(* Logix 5000 project; controller MV vendor 1 type 14 code 217 rev 31.11; software revision 31.00; part 28 of 53 *)
(* tags used below, declared in another part *)
   active : BOOL;
   CWD : CHECKWORD_FLAGS;
   FVHR18_2505 : PlantItem;   // Valve FVHR18_25/05
   FVHR18_2506 : PlantItem;   // Valve FVHR18_25/06
   FVHR26_3101 : PlantItem;   // Valve FVHR26_31/01
   FVHR26_3102 : PlantItem;   // Valve FVHR26_31/02
   FVHR26_3103 : PlantItem;   // Valve FVHR26_31/03
   FVHRCH201 : PlantItem;   // Valve FVHRCH201
   FVHRCH202 : PlantItem;   // Valve FVHRCH202
   FVHRCW01 : PlantItem;   // Valve FVHRCW01
   FVHRM01 : PlantItem;   // Valve FVHRM01
   FVHRM02 : PlantItem;   // Valve FVHRM02
   FVHRM03 : PlantItem;   // Valve FVHRM03
   FVHRM04 : PlantItem;   // Valve FVHRM04
   FVHRMD01 : PlantItem;   // Valve FVHRMD01
   IGI_TestBit : BOOL;
   MC_B243 : INT[255];   // CH2 ROUTE Channel 2 route requ est flags
   MC_CD_T1 : PlantItem;   // CD_T1
   MC_CH2_CIP_BYPASS_Conditions : BOOL;
   MC_CH2_CIP_BYPASS_DrainConditions : BOOL;
   MC_CH2_CIP_Messages : STRING[20];   // CH2 CIP Scada Messages
   MC_CH2_CIP_YST_Scb_Bypass : BOOL;
   MC_CH2_FVBYPASS_H2O_Flush : BOOL;
   MC_CIP_CH2_Strings_HopRinse : STRING[30];
   MC_CIP_String_Result : DINT;
   MC_FL_D1 : PlantItem;   // FL_D1
   MC_N10 : INT[255];   // SETTINGS
   MC_N100 : INT[255];   // C1_PLC Channel 1 PLC data
   MC_N104 : INT[255];   // CH1 REPORT Channel 1 CIP report file
   MC_N120 : INT[255];   // C2 PLC Channel 2 PLC data
   MC_N122 : INT[255];   // CH2 PROG Channel 2 CIP progra m
   MC_N124 : INT[255];   // CH2 REPORT Channel 2 CIP report file
   MC_N200 : INT[255];   // CHK_WORK Plant item fault che cking work area
   MC_N7 : INT[255];   // INTEGER
   MC_N80 : INT[255];   // SRV1_PLC Detergent tank 1 ser vice PLC data
   MC_N80_19_0_Storagebit : BOOL;
   MC_N81 : INT[255];   // SV1_PC Detergent tank 1 ser vice PC to PLC data
   MC_P3 : PlantItem;   // P3
   MC_SFile : INT[255];   // SLC Equivalent System File, So Original Code Can Remain
   MC_SV1 : PlantItem;   // SV1
   MC_T125 : TIMER[255];   // CH2 TIMERS Channel 2 timers
   MC_T4 : TIMER[255];   // TIMER
   MC_T85 : TIMER[255];   // SV1 TIMERS Detergent tank 1 ser vice timers
(* MC_Common, continued *)

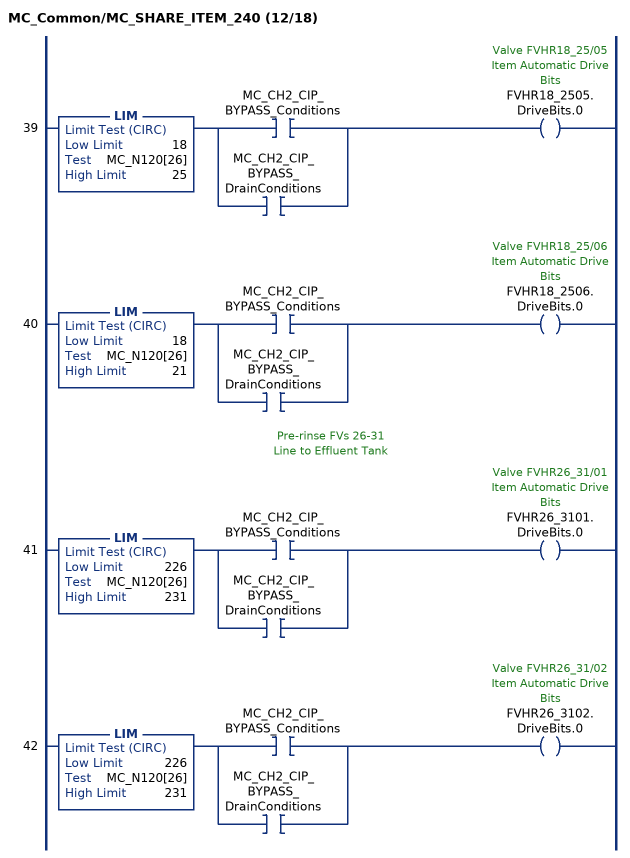
   [picture p556: MC_Common/MC_SHARE_ITEM_240 rungs 39-42]
   39: LIM(18,MC_N120[26],25)[XIC(MC_CH2_CIP_BYPASS_Conditions) ,XIC(MC_CH2_CIP_BYPASS_DrainConditions) ]OTE(FVHR18_2505.DriveBits.0);
   40: LIM(18,MC_N120[26],21)[XIC(MC_CH2_CIP_BYPASS_Conditions) ,XIC(MC_CH2_CIP_BYPASS_DrainConditions) ]OTE(FVHR18_2506.DriveBits.0);
   // Pre-rinse FVs 26-31
   // Line to Effluent Tank
   41: LIM(226,MC_N120[26],231)[XIC(MC_CH2_CIP_BYPASS_Conditions) ,XIC(MC_CH2_CIP_BYPASS_DrainConditions) ]OTE(FVHR26_3101.DriveBits.0);
   42: LIM(226,MC_N120[26],231)[XIC(MC_CH2_CIP_BYPASS_Conditions) ,XIC(MC_CH2_CIP_BYPASS_DrainConditions) ]OTE(FVHR26_3102.DriveBits.0);
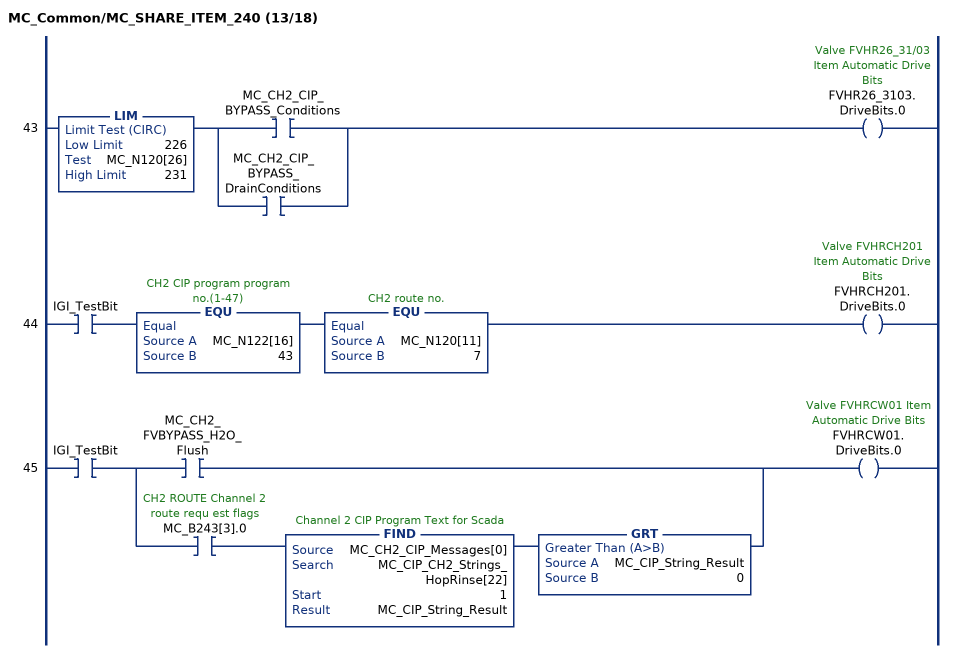
   43: LIM(226,MC_N120[26],231)[XIC(MC_CH2_CIP_BYPASS_Conditions) ,XIC(MC_CH2_CIP_BYPASS_DrainConditions) ]OTE(FVHR26_3103.DriveBits.0);
   44: XIC(IGI_TestBit)EQU(MC_N122[16],43)EQU(MC_N120[11],7)OTE(FVHRCH201.DriveBits.0);
   45: XIC(IGI_TestBit)[XIC(MC_CH2_FVBYPASS_H2O_Flush) ,XIC(MC_B243[3].0) FIND(MC_CH2_CIP_Messages[0],MC_CIP_CH2_Strings_HopRinse[22],1,MC_CIP_String_Result) GRT(MC_CIP_String_Result,0) ]OTE(FVHRCW01.DriveBits.0);
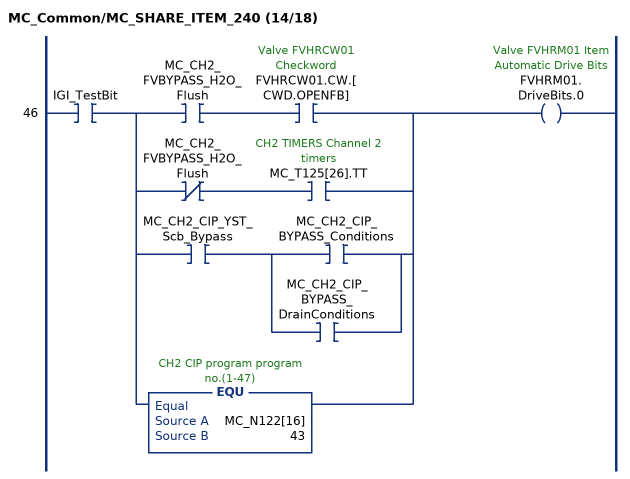
   46: XIC(IGI_TestBit)[XIC(MC_CH2_FVBYPASS_H2O_Flush) XIC(FVHRCW01.CW.[CWD.OPENFB]) ,XIO(MC_CH2_FVBYPASS_H2O_Flush) XIC(MC_T125[26].TT) ,XIC(MC_CH2_CIP_YST_Scb_Bypass) [XIC(MC_CH2_CIP_BYPASS_Conditions) ,XIC(MC_CH2_CIP_BYPASS_DrainConditions) ] ,EQU(MC_N122[16],43) ]OTE(FVHRM01.DriveBits.0);
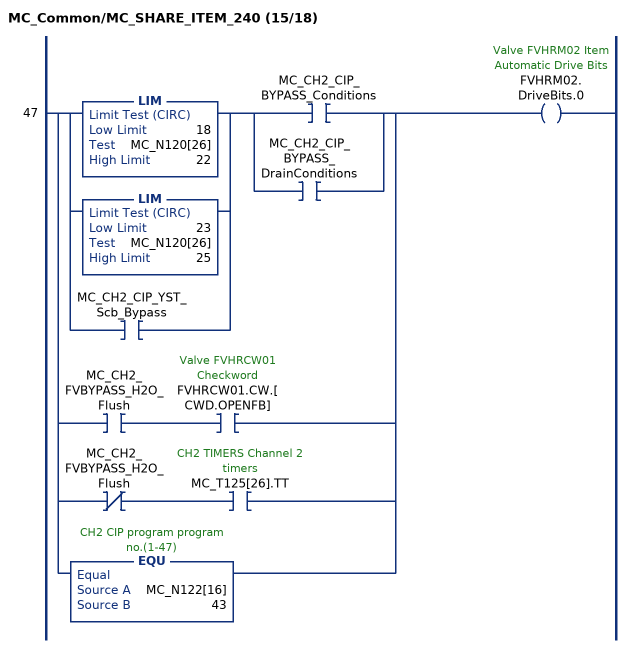
   47: [[LIM(18,MC_N120[26],22) ,LIM(23,MC_N120[26],25) ,XIC(MC_CH2_CIP_YST_Scb_Bypass) ] [XIC(MC_CH2_CIP_BYPASS_Conditions) ,XIC(MC_CH2_CIP_BYPASS_DrainConditions) ] ,XIC(MC_CH2_FVBYPASS_H2O_Flush) XIC(FVHRCW01.CW.[CWD.OPENFB]) ,XIO(MC_CH2_FVBYPASS_H2O_Flush) XIC(MC_T125[26].TT) ,EQU(MC_N122[16],43) ]OTE(FVHRM02.DriveBits.0);
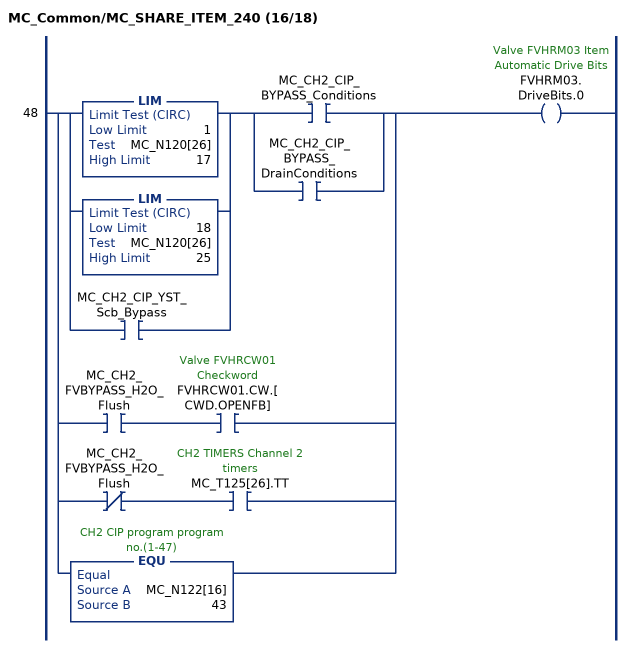
   48: [[LIM(1,MC_N120[26],17) ,LIM(18,MC_N120[26],25) ,XIC(MC_CH2_CIP_YST_Scb_Bypass) ] [XIC(MC_CH2_CIP_BYPASS_Conditions) ,XIC(MC_CH2_CIP_BYPASS_DrainConditions) ] ,XIC(MC_CH2_FVBYPASS_H2O_Flush) XIC(FVHRCW01.CW.[CWD.OPENFB]) ,XIO(MC_CH2_FVBYPASS_H2O_Flush) XIC(MC_T125[26].TT) ,EQU(MC_N122[16],43) ]OTE(FVHRM03.DriveBits.0);
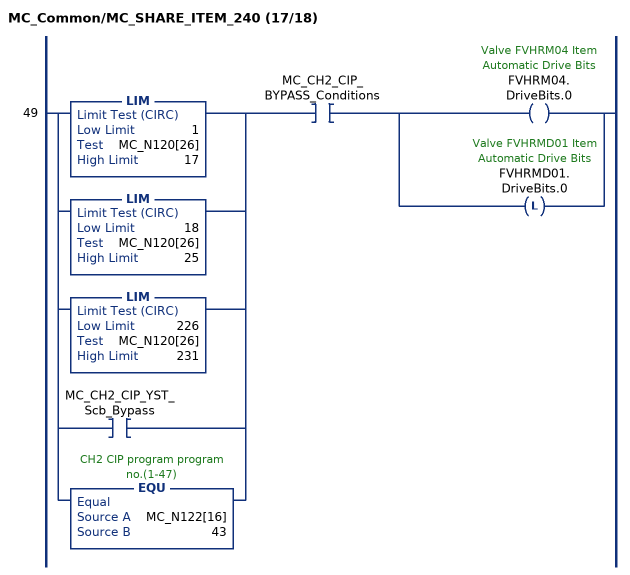
   49: [LIM(1,MC_N120[26],17) ,LIM(18,MC_N120[26],25) ,LIM(226,MC_N120[26],231) ,XIC(MC_CH2_CIP_YST_Scb_Bypass) ,EQU(MC_N122[16],43) ]XIC(MC_CH2_CIP_BYPASS_Conditions)[OTE(FVHRM04.DriveBits.0) ,OTL(FVHRMD01.DriveBits.0) ];
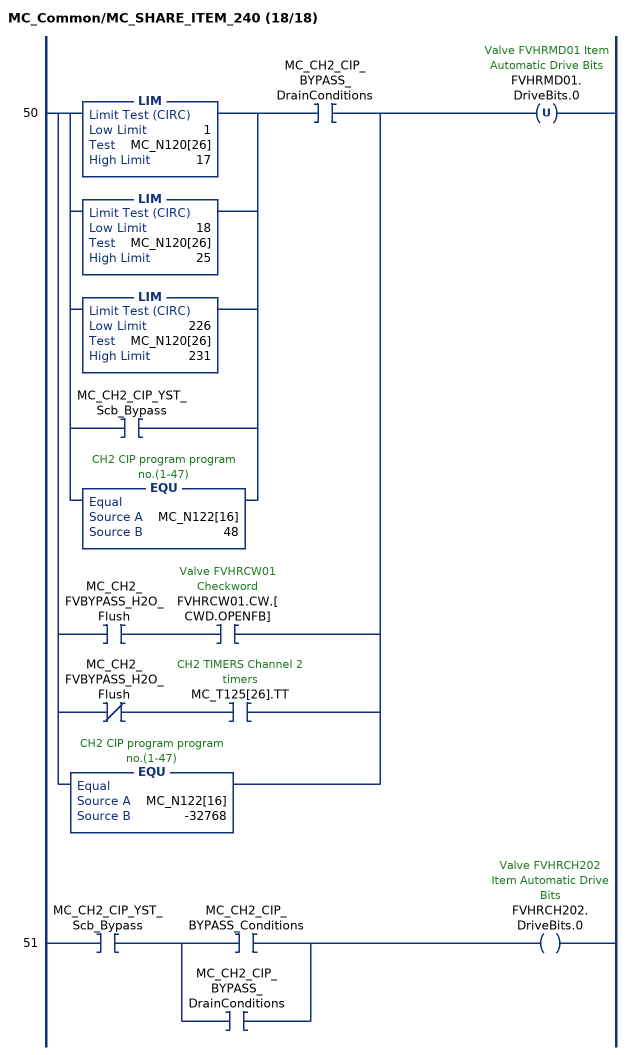
   50: [[LIM(1,MC_N120[26],17) ,LIM(18,MC_N120[26],25) ,LIM(226,MC_N120[26],231) ,XIC(MC_CH2_CIP_YST_Scb_Bypass) ,EQU(MC_N122[16],48) ] XIC(MC_CH2_CIP_BYPASS_DrainConditions) ,XIC(MC_CH2_FVBYPASS_H2O_Flush) XIC(FVHRCW01.CW.[CWD.OPENFB]) ,XIO(MC_CH2_FVBYPASS_H2O_Flush) XIC(MC_T125[26].TT) ,EQU(MC_N122[16],-32768) ]OTU(FVHRMD01.DriveBits.0);
   51: XIC(MC_CH2_CIP_YST_Scb_Bypass)[XIC(MC_CH2_CIP_BYPASS_Conditions) ,XIC(MC_CH2_CIP_BYPASS_DrainConditions) ]OTE(FVHRCH202.DriveBits.0);
END_ROUTINE

ROUTINE MC_SRV1_CMD_81   (* ladder *)
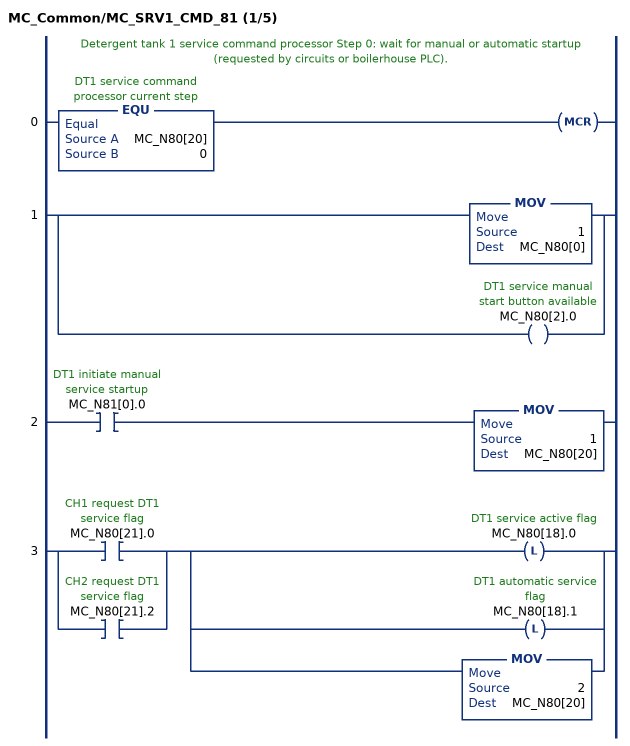
   // Detergent tank 1 service command processor Step 0: wait for manual or automatic startup (requested by circuits or boilerhouse PLC).
   0: EQU(MC_N80[20],0)MCR();
   1: [MOV(1,MC_N80[0]) ,OTE(MC_N80[2].0) ];
   2: XIC(MC_N81[0].0)MOV(1,MC_N80[20]);
   3: [XIC(MC_N80[21].0) ,XIC(MC_N80[21].2) ][OTL(MC_N80[18].0) ,OTL(MC_N80[18].1) ,MOV(2,MC_N80[20]) ];
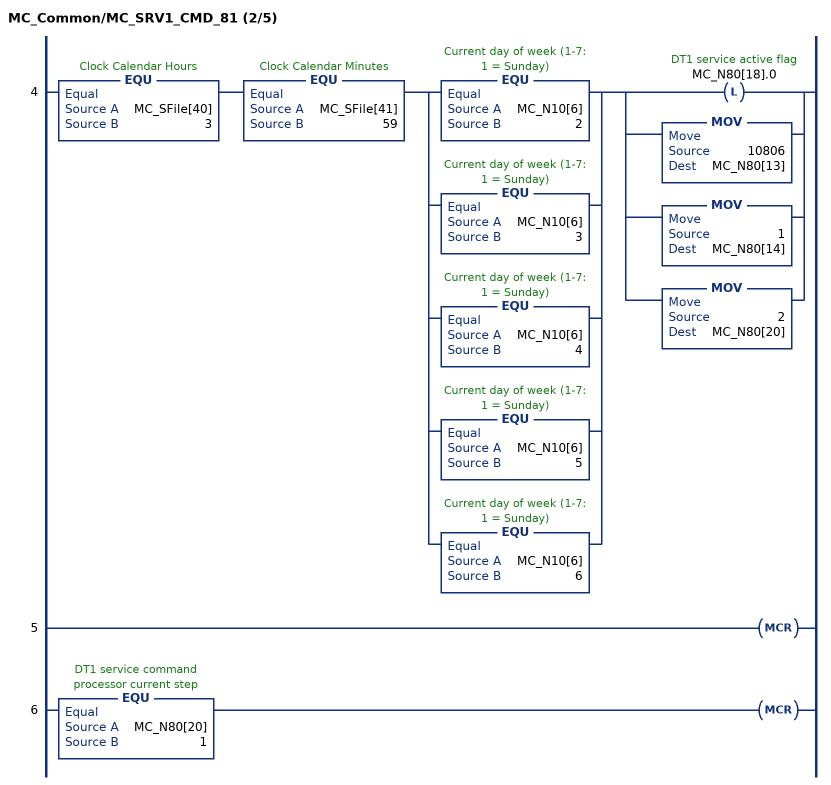
   4: EQU(MC_SFile[40],3)EQU(MC_SFile[41],59)[EQU(MC_N10[6],2) ,EQU(MC_N10[6],3) ,EQU(MC_N10[6],4) ,EQU(MC_N10[6],5) ,EQU(MC_N10[6],6) ][OTL(MC_N80[18].0) ,MOV(10806,MC_N80[13]) ,MOV(1,MC_N80[14]) ,MOV(2,MC_N80[20]) ];
   5: MCR();
   6: EQU(MC_N80[20],1)MCR();
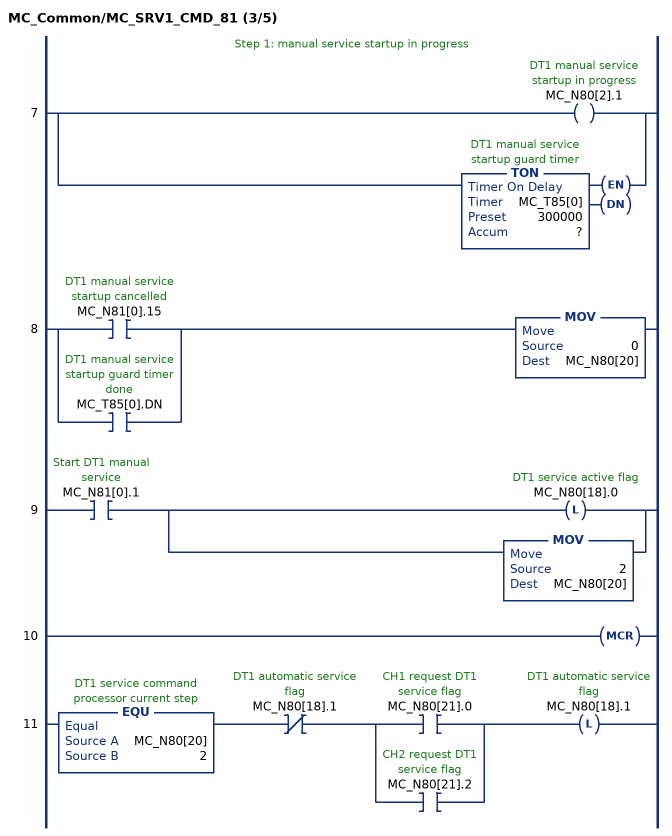
   // Step 1: manual service startup in progress
   7: [OTE(MC_N80[2].1) ,TON(MC_T85[0],?,?) ];
   8: [XIC(MC_N81[0].15) ,XIC(MC_T85[0].DN) ]MOV(0,MC_N80[20]);
   9: XIC(MC_N81[0].1)[OTL(MC_N80[18].0) ,MOV(2,MC_N80[20]) ];
   10: MCR();
   11: EQU(MC_N80[20],2)XIO(MC_N80[18].1)[XIC(MC_N80[21].0) ,XIC(MC_N80[21].2) ]OTL(MC_N80[18].1);
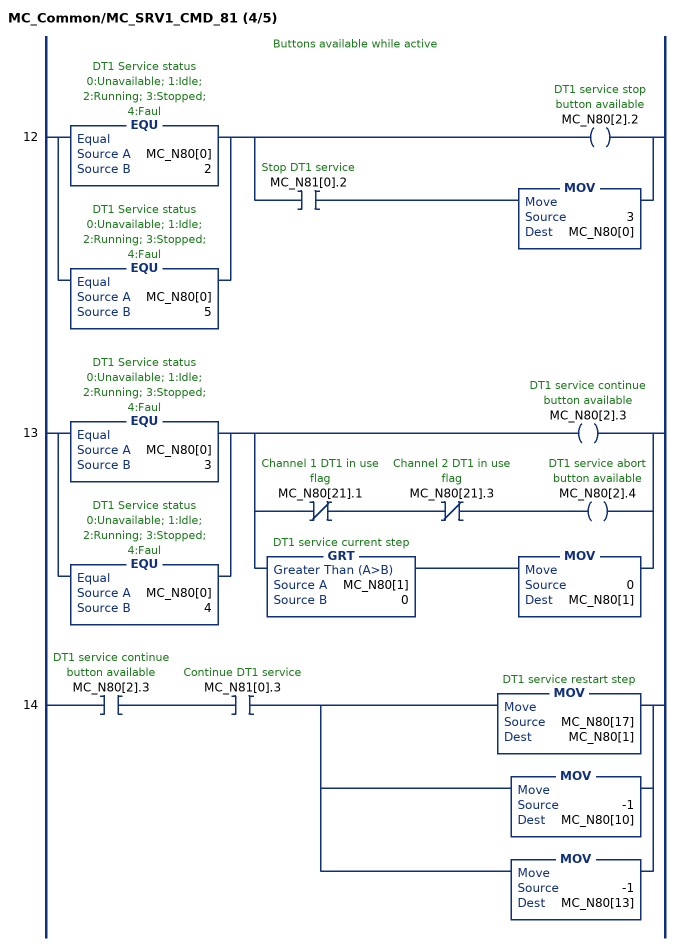
   // Buttons available while active
   12: [EQU(MC_N80[0],2) ,EQU(MC_N80[0],5) ][OTE(MC_N80[2].2) ,XIC(MC_N81[0].2) MOV(3,MC_N80[0]) ];
   13: [EQU(MC_N80[0],3) ,EQU(MC_N80[0],4) ][OTE(MC_N80[2].3) ,XIO(MC_N80[21].1) XIO(MC_N80[21].3) OTE(MC_N80[2].4) ,GRT(MC_N80[1],0) MOV(0,MC_N80[1]) ];
   14: XIC(MC_N80[2].3)XIC(MC_N81[0].3)[MOV(MC_N80[17],MC_N80[1]) ,MOV(-1,MC_N80[10]) ,MOV(-1,MC_N80[13]) ];
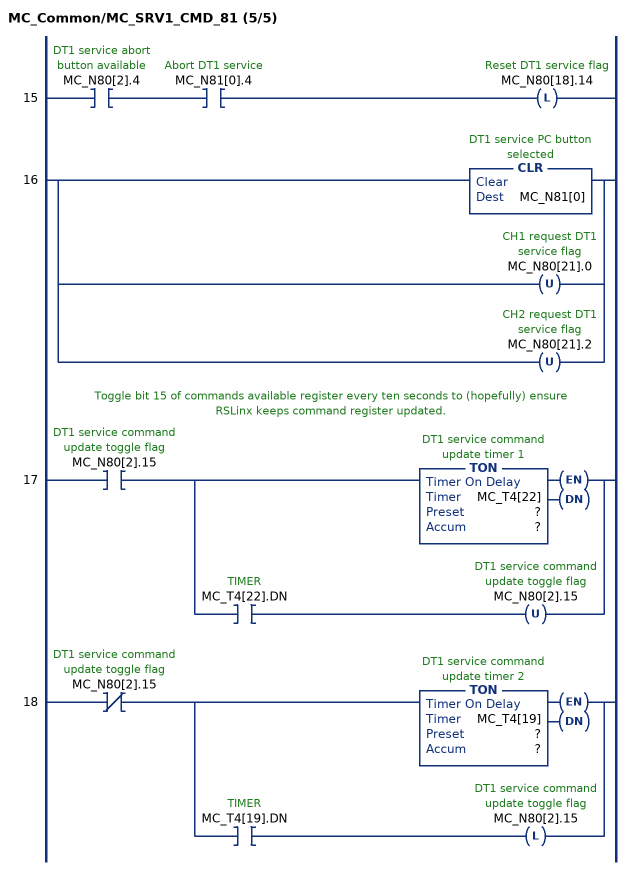
   15: XIC(MC_N80[2].4)XIC(MC_N81[0].4)OTL(MC_N80[18].14);
   16: [CLR(MC_N81[0]) ,OTU(MC_N80[21].0) ,OTU(MC_N80[21].2) ];
   // Toggle bit 15 of commands available register every ten seconds to (hopefully) ensure RSLinx keeps command register updated.
   17: XIC(MC_N80[2].15)[TON(MC_T4[22],?,?) ,XIC(MC_T4[22].DN) OTU(MC_N80[2].15) ];
   18: XIO(MC_N80[2].15)[TON(MC_T4[19],?,?) ,XIC(MC_T4[19].DN) OTL(MC_N80[2].15) ];
END_ROUTINE

ROUTINE MC_SRV1_MCP_80   (* ladder *)
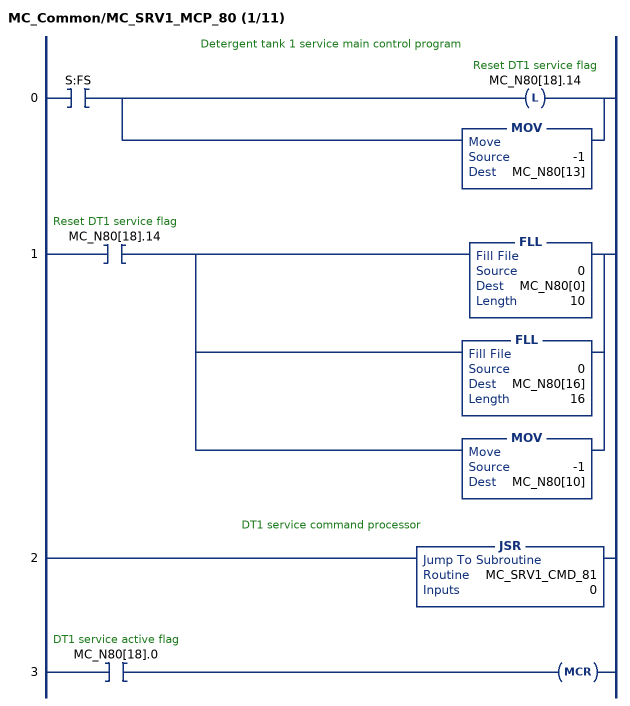
   // Detergent tank 1 service main control program
   0: XIC(S:FS)[OTL(MC_N80[18].14) ,MOV(-1,MC_N80[13]) ];
   1: XIC(MC_N80[18].14)[FLL(0,MC_N80[0],10) ,FLL(0,MC_N80[16],16) ,MOV(-1,MC_N80[10]) ];
   // DT1 service command processor
   2: JSR(MC_SRV1_CMD_81,0);
   3: XIC(MC_N80[18].0)MCR();
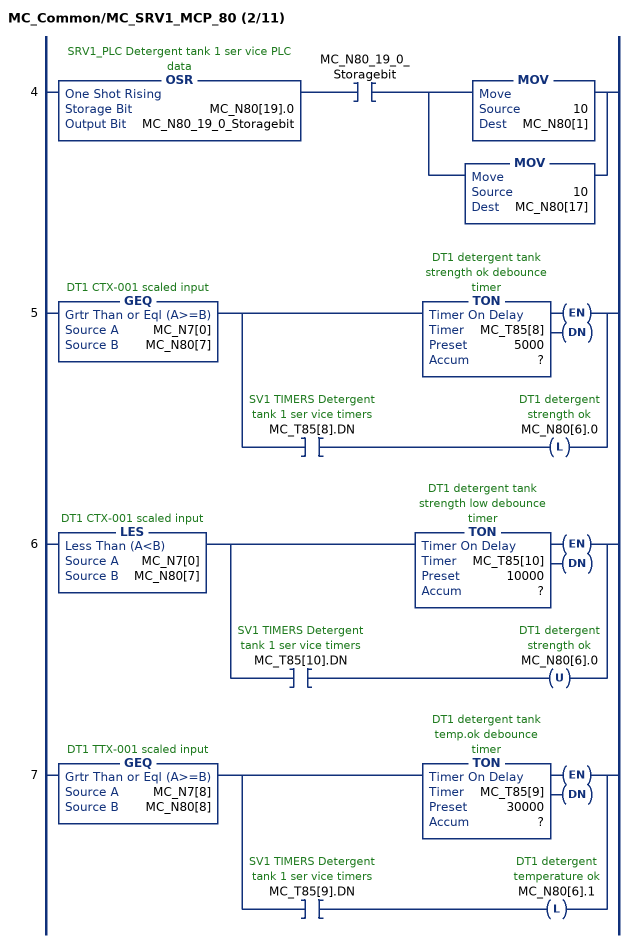
   4: OSR(MC_N80[19].0,MC_N80_19_0_Storagebit)XIC(MC_N80_19_0_Storagebit)[MOV(10,MC_N80[1]) ,MOV(10,MC_N80[17]) ];
   5: GEQ(MC_N7[0],MC_N80[7])[TON(MC_T85[8],?,?) ,XIC(MC_T85[8].DN) OTL(MC_N80[6].0) ];
   6: LES(MC_N7[0],MC_N80[7])[TON(MC_T85[10],?,?) ,XIC(MC_T85[10].DN) OTU(MC_N80[6].0) ];
   7: GEQ(MC_N7[8],MC_N80[8])[TON(MC_T85[9],?,?) ,XIC(MC_T85[9].DN) OTL(MC_N80[6].1) ];
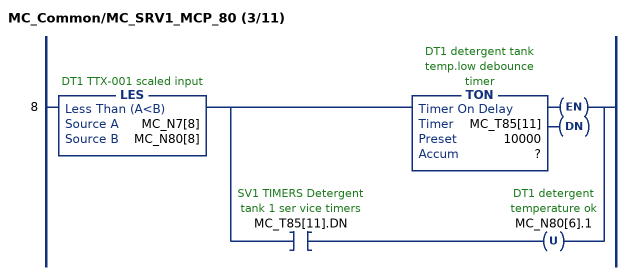
   8: LES(MC_N7[8],MC_N80[8])[TON(MC_T85[11],?,?) ,XIC(MC_T85[11].DN) OTU(MC_N80[6].1) ];
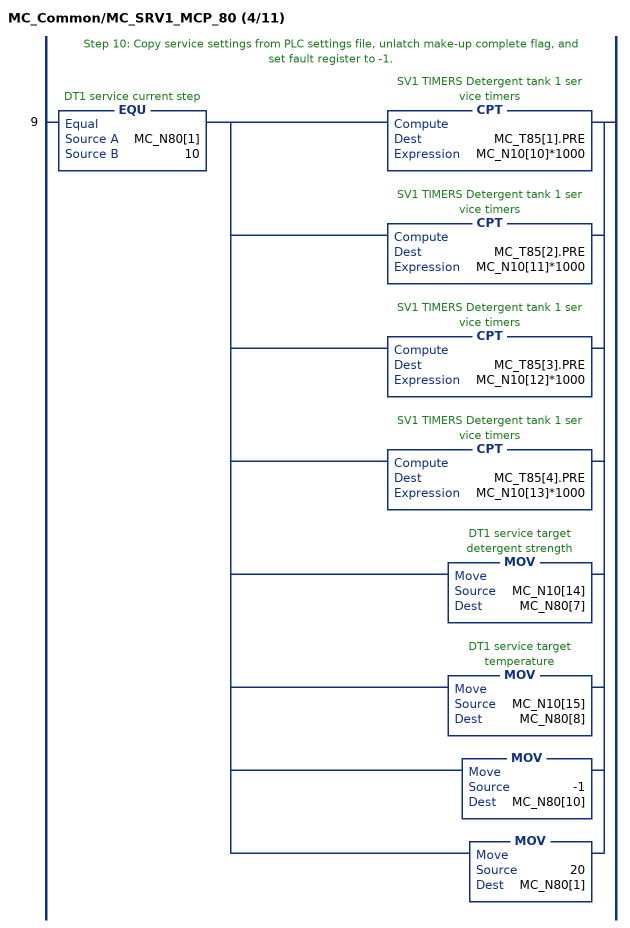
   // Step 10: Copy service settings from PLC settings file, unlatch make-up complete flag, and set fault register to -1.
   9: EQU(MC_N80[1],10)[CPT(MC_T85[1].PRE,MC_N10[10]*1000) ,CPT(MC_T85[2].PRE,MC_N10[11]*1000) ,CPT(MC_T85[3].PRE,MC_N10[12]*1000) ,CPT(MC_T85[4].PRE,MC_N10[13]*1000) ,MOV(MC_N10[14],MC_N80[7]) ,MOV(MC_N10[15],MC_N80[8]) ,MOV(-1,MC_N80[10]) ,MOV(20,MC_N80[1]) ];
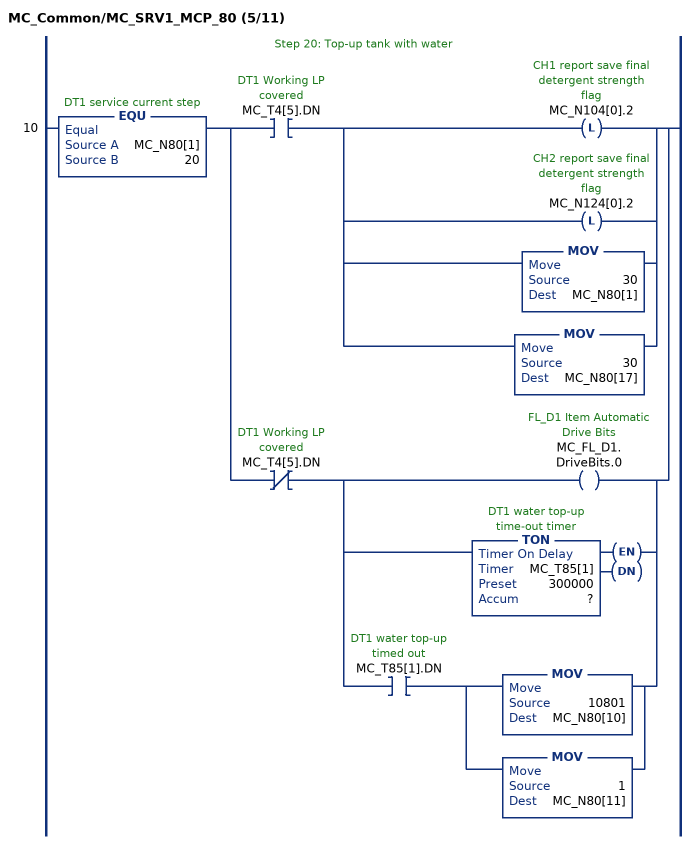
   // Step 20: Top-up tank with water
   10: EQU(MC_N80[1],20)[XIC(MC_T4[5].DN) [OTL(MC_N104[0].2) ,OTL(MC_N124[0].2) ,MOV(30,MC_N80[1]) ,MOV(30,MC_N80[17]) ] ,XIO(MC_T4[5].DN) [OTE(MC_FL_D1.DriveBits.0) ,TON(MC_T85[1],?,?) ,XIC(MC_T85[1].DN) [MOV(10801,MC_N80[10]) ,MOV(1,MC_N80[11]) ] ] ];
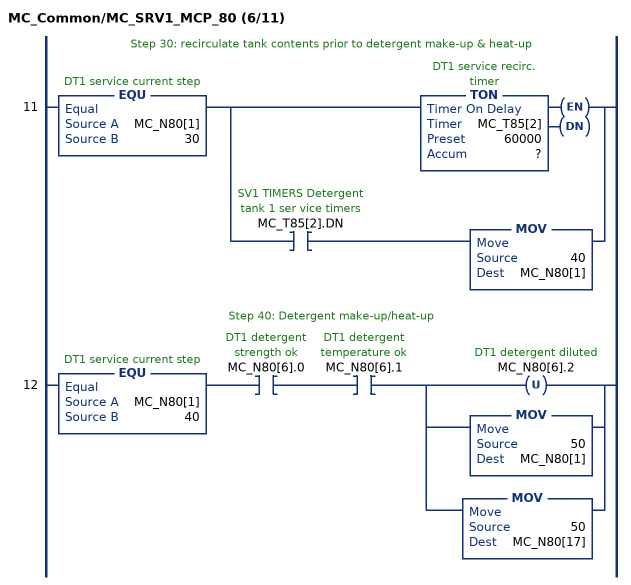
   // Step 30: recirculate tank contents prior to detergent make-up & heat-up
   11: EQU(MC_N80[1],30)[TON(MC_T85[2],?,?) ,XIC(MC_T85[2].DN) MOV(40,MC_N80[1]) ];
   // Step 40: Detergent make-up/heat-up
   12: EQU(MC_N80[1],40)XIC(MC_N80[6].0)XIC(MC_N80[6].1)[OTU(MC_N80[6].2) ,MOV(50,MC_N80[1]) ,MOV(50,MC_N80[17]) ];
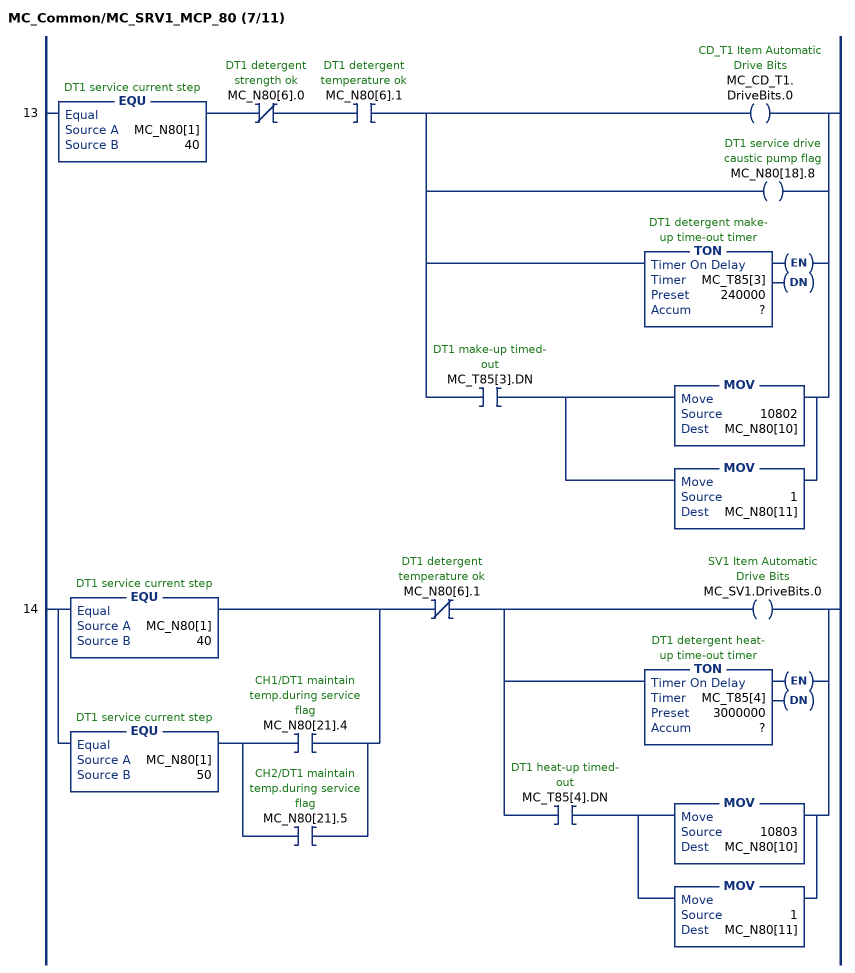
   13: EQU(MC_N80[1],40)XIO(MC_N80[6].0)XIC(MC_N80[6].1)[[OTE(MC_CD_T1.DriveBits.0) ,OTE(MC_N80[18].8) ] ,TON(MC_T85[3],?,?) ,XIC(MC_T85[3].DN) [MOV(10802,MC_N80[10]) ,MOV(1,MC_N80[11]) ] ];
   14: [EQU(MC_N80[1],40) ,EQU(MC_N80[1],50) [XIC(MC_N80[21].4) ,XIC(MC_N80[21].5) ] ]XIO(MC_N80[6].1)[OTE(MC_SV1.DriveBits.0) ,TON(MC_T85[4],?,?) ,XIC(MC_T85[4].DN) [MOV(10803,MC_N80[10]) ,MOV(1,MC_N80[11]) ] ];
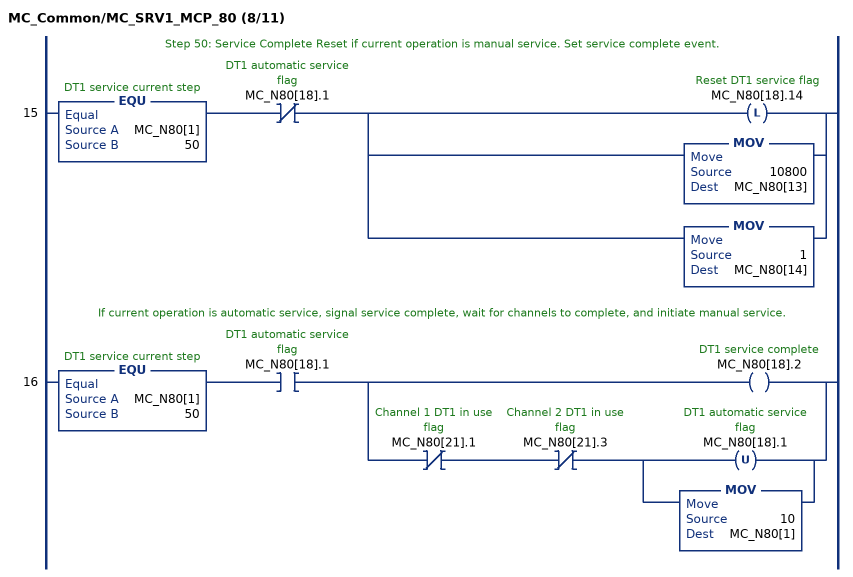
   // Step 50: Service Complete Reset if current operation is manual service. Set service complete event.
   15: EQU(MC_N80[1],50)XIO(MC_N80[18].1)[OTL(MC_N80[18].14) ,MOV(10800,MC_N80[13]) ,MOV(1,MC_N80[14]) ];
   // If current operation is automatic service, signal service complete, wait for channels to complete, and initiate manual service.
   16: EQU(MC_N80[1],50)XIC(MC_N80[18].1)[OTE(MC_N80[18].2) ,XIO(MC_N80[21].1) XIO(MC_N80[21].3) [OTU(MC_N80[18].1) ,MOV(10,MC_N80[1]) ] ];
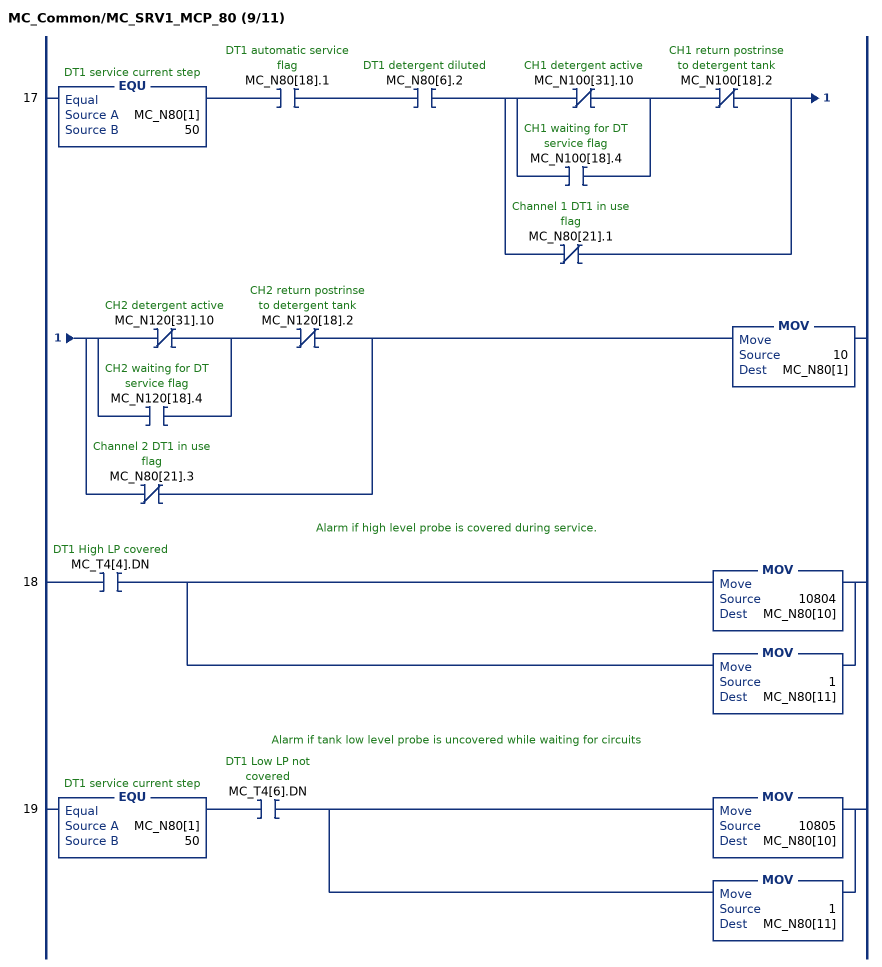
   17: EQU(MC_N80[1],50)XIC(MC_N80[18].1)XIC(MC_N80[6].2)[[XIO(MC_N100[31].10) ,XIC(MC_N100[18].4) ] XIO(MC_N100[18].2) ,XIO(MC_N80[21].1) ][[XIO(MC_N120[31].10) ,XIC(MC_N120[18].4) ] XIO(MC_N120[18].2) ,XIO(MC_N80[21].3) ]MOV(10,MC_N80[1]);
   // Alarm if high level probe is covered during service.
   18: XIC(MC_T4[4].DN)[MOV(10804,MC_N80[10]) ,MOV(1,MC_N80[11]) ];
   // Alarm if tank low level probe is uncovered while waiting for circuits
   19: EQU(MC_N80[1],50)XIC(MC_T4[6].DN)[MOV(10805,MC_N80[10]) ,MOV(1,MC_N80[11]) ];
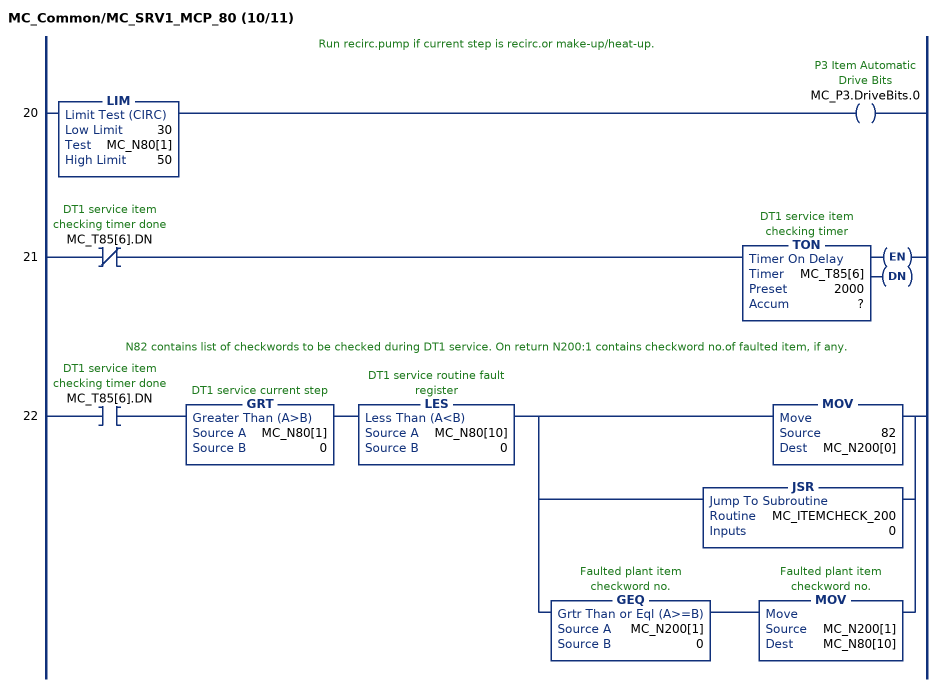
   // Run recirc.pump if current step is recirc.or make-up/heat-up.
   20: LIM(30,MC_N80[1],50)OTE(MC_P3.DriveBits.0);
   21: XIO(MC_T85[6].DN)TON(MC_T85[6],?,?);
   // N82 contains list of checkwords to be checked during DT1 service. On return N200:1 contains checkword no.of faulted item, if any.
   22: XIC(MC_T85[6].DN)GRT(MC_N80[1],0)LES(MC_N80[10],0)[MOV(82,MC_N200[0]) ,JSR(MC_ITEMCHECK_200,0) ,GEQ(MC_N200[1],0) MOV(MC_N200[1],MC_N80[10]) ];
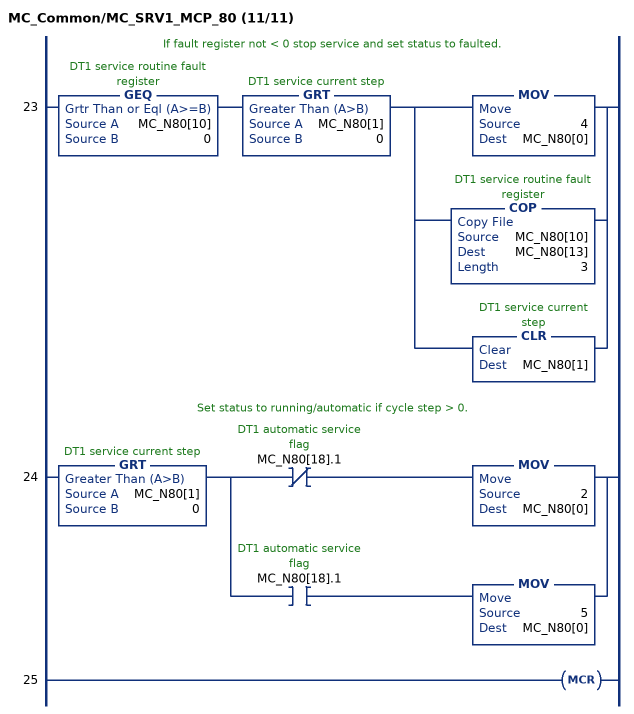
   // If fault register not < 0 stop service and set status to faulted.
   23: GEQ(MC_N80[10],0)GRT(MC_N80[1],0)[MOV(4,MC_N80[0]) ,COP(MC_N80[10],MC_N80[13],3) ,CLR(MC_N80[1]) ];
   // Set status to running/automatic if cycle step > 0.
   24: GRT(MC_N80[1],0)[XIO(MC_N80[18].1) MOV(2,MC_N80[0]) ,XIC(MC_N80[18].1) MOV(5,MC_N80[0]) ];
   25: MCR();
END_ROUTINE
